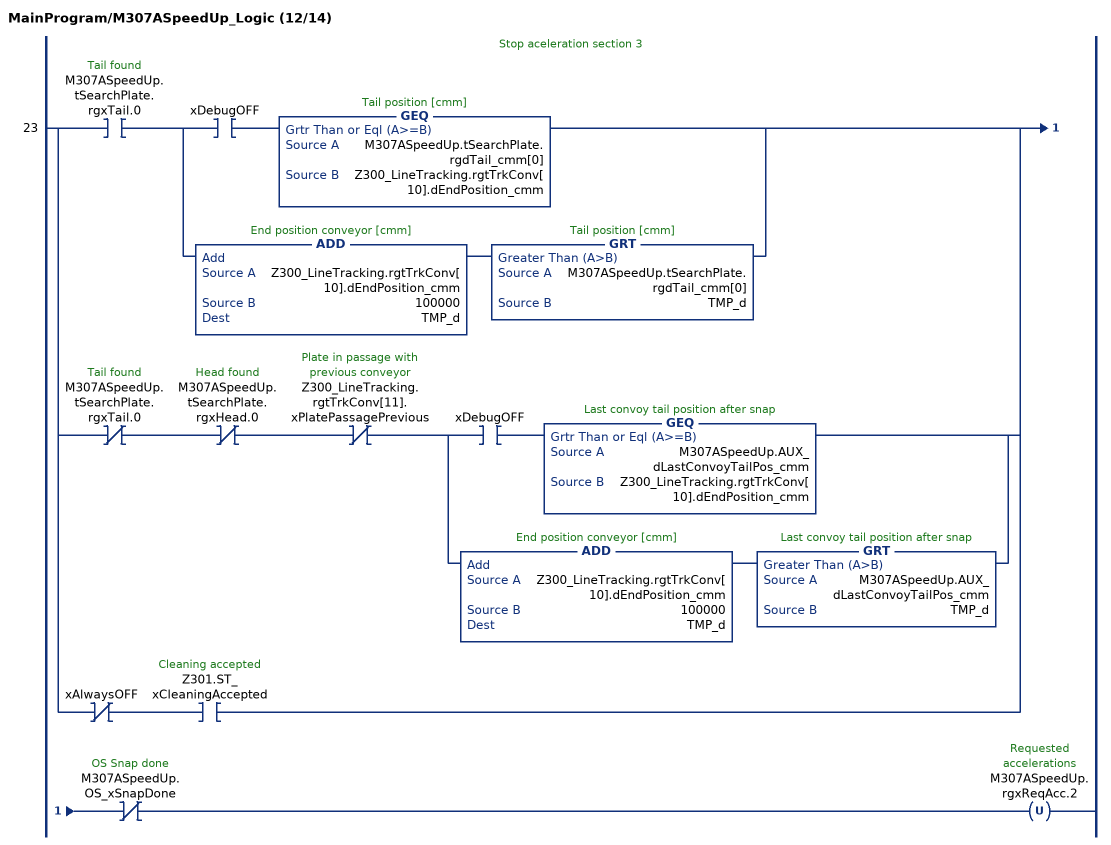
   // Stop aceleration section 3
   23: [XIC(M307ASpeedUp.tSearchPlate.rgxTail.0) [XIC(xDebugOFF) GEQ(M307ASpeedUp.tSearchPlate.rgdTail_cmm[0],Z300_LineTracking.rgtTrkConv[10].dEndPosition_cmm) ,ADD(Z300_LineTracking.rgtTrkConv[10].dEndPosition_cmm,100000,TMP_d) GRT(M307ASpeedUp.tSearchPlate.rgdTail_cmm[0],TMP_d) ] ,XIO(M307ASpeedUp.tSearchPlate.rgxTail.0) XIO(M307ASpeedUp.tSearchPlate.rgxHead.0) XIO(Z300_LineTracking.rgtTrkConv[11].xPlatePassagePrevious) [XIC(xDebugOFF) GEQ(M307ASpeedUp.AUX_dLastConvoyTailPos_cmm,Z300_LineTracking.rgtTrkConv[10].dEndPosition_cmm) ,ADD(Z300_LineTracking.rgtTrkConv[10].dEndPosition_cmm,100000,TMP_d) GRT(M307ASpeedUp.AUX_dLastConvoyTailPos_cmm,TMP_d) ] ,XIO(xAlwaysOFF) XIC(Z301.ST_xCleaningAccepted) ]XIO(M307ASpeedUp.OS_xSnapDone)OTU(M307ASpeedUp.rgxReqAcc.2);
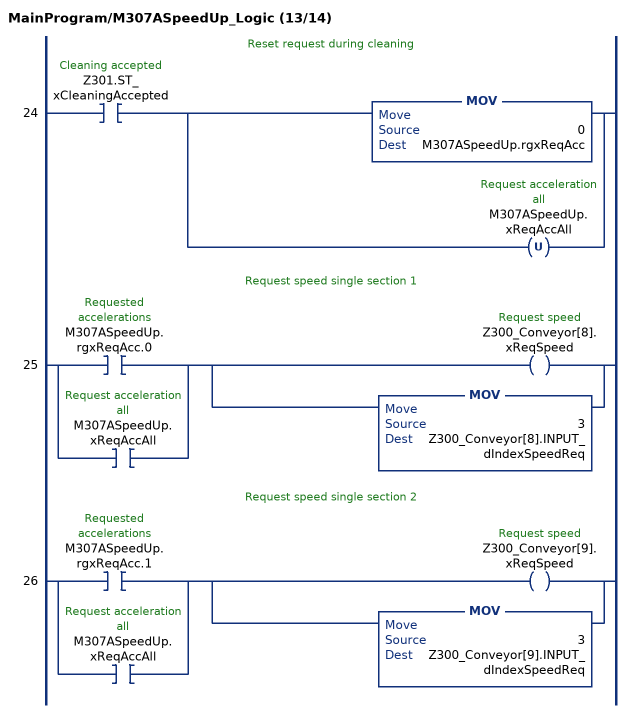
   // Reset request during cleaning
   24: XIC(Z301.ST_xCleaningAccepted)[MOV(0,M307ASpeedUp.rgxReqAcc) ,OTU(M307ASpeedUp.xReqAccAll) ];
   // Request speed single section 1
   25: [XIC(M307ASpeedUp.rgxReqAcc.0) ,XIC(M307ASpeedUp.xReqAccAll) ][OTE(Z300_Conveyor[8].xReqSpeed) ,MOV(3,Z300_Conveyor[8].INPUT_dIndexSpeedReq) ];
   // Request speed single section 2
   26: [XIC(M307ASpeedUp.rgxReqAcc.1) ,XIC(M307ASpeedUp.xReqAccAll) ][OTE(Z300_Conveyor[9].xReqSpeed) ,MOV(3,Z300_Conveyor[9].INPUT_dIndexSpeedReq) ];
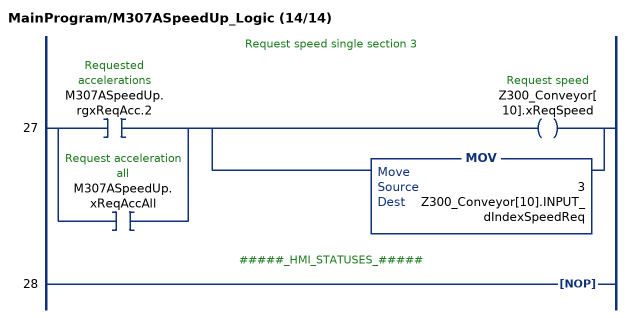
   // Request speed single section 3
   27: [XIC(M307ASpeedUp.rgxReqAcc.2) ,XIC(M307ASpeedUp.xReqAccAll) ][OTE(Z300_Conveyor[10].xReqSpeed) ,MOV(3,Z300_Conveyor[10].INPUT_dIndexSpeedReq) ];
   // #####_HMI_STATUSES_#####
   28: NOP();
END_ROUTINE

ROUTINE M30xTrimDeck_Faults   (* ladder *)
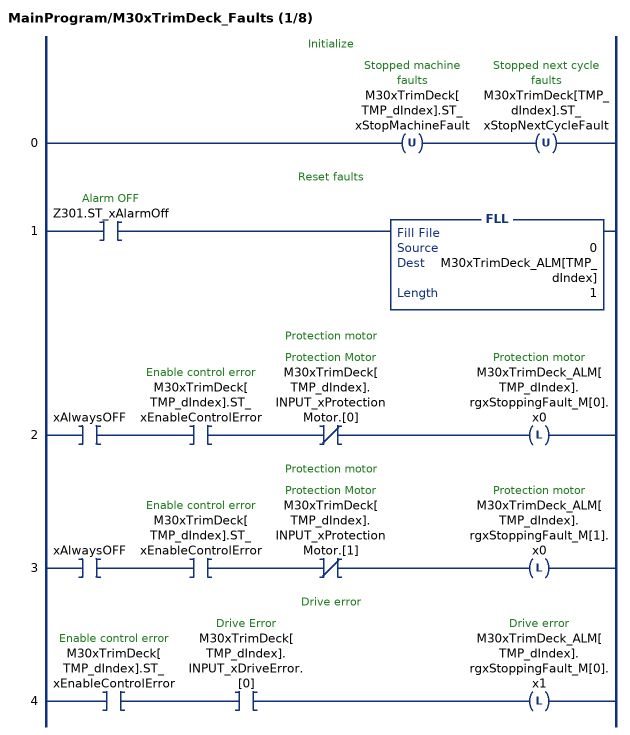
   // Initialize
   0: OTU(M30xTrimDeck[TMP_dIndex].ST_xStopMachineFault)OTU(M30xTrimDeck[TMP_dIndex].ST_xStopNextCycleFault);
   // Reset faults
   1: XIC(Z301.ST_xAlarmOff)FLL(0,M30xTrimDeck_ALM[TMP_dIndex],1);
   // Protection motor
   2: XIC(xAlwaysOFF)XIC(M30xTrimDeck[TMP_dIndex].ST_xEnableControlError)XIO(M30xTrimDeck[TMP_dIndex].INPUT_xProtectionMotor.[0])OTL(M30xTrimDeck_ALM[TMP_dIndex].rgxStoppingFault_M[0].x0);
   // Protection motor
   3: XIC(xAlwaysOFF)XIC(M30xTrimDeck[TMP_dIndex].ST_xEnableControlError)XIO(M30xTrimDeck[TMP_dIndex].INPUT_xProtectionMotor.[1])OTL(M30xTrimDeck_ALM[TMP_dIndex].rgxStoppingFault_M[1].x0);
   // Drive error
   4: XIC(M30xTrimDeck[TMP_dIndex].ST_xEnableControlError)XIC(M30xTrimDeck[TMP_dIndex].INPUT_xDriveError.[0])OTL(M30xTrimDeck_ALM[TMP_dIndex].rgxStoppingFault_M[0].x1);
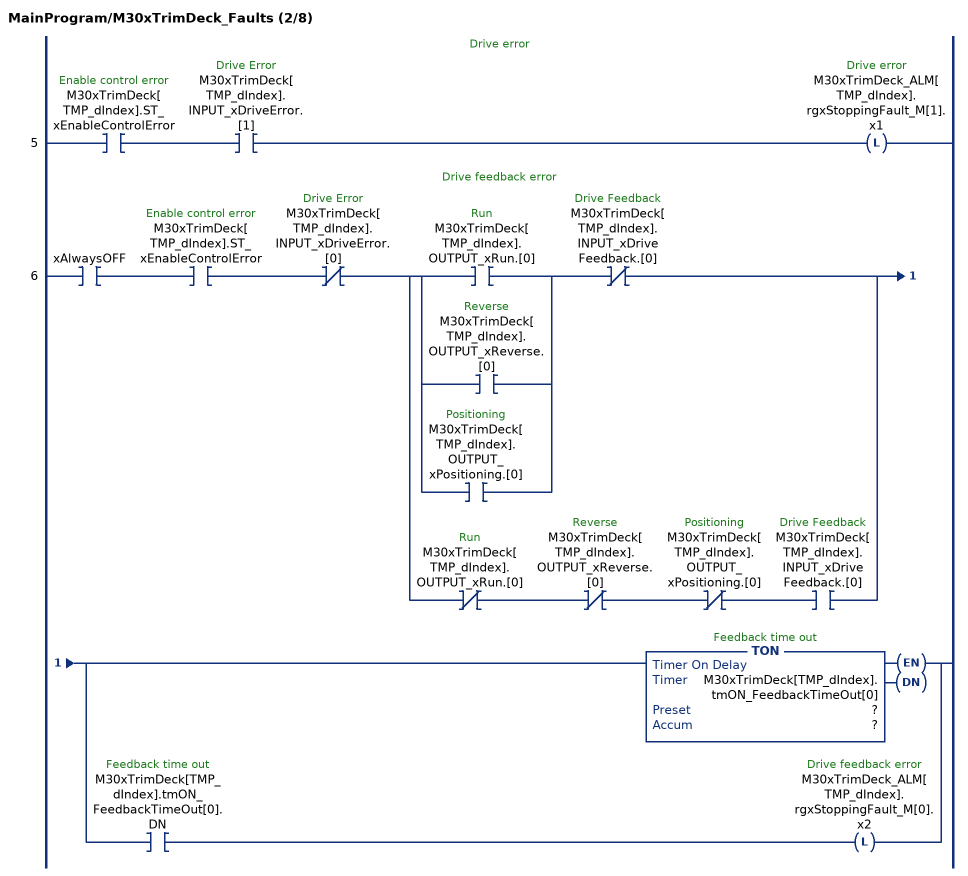
   // Drive error
   5: XIC(M30xTrimDeck[TMP_dIndex].ST_xEnableControlError)XIC(M30xTrimDeck[TMP_dIndex].INPUT_xDriveError.[1])OTL(M30xTrimDeck_ALM[TMP_dIndex].rgxStoppingFault_M[1].x1);
   // Drive feedback error
   6: XIC(xAlwaysOFF)XIC(M30xTrimDeck[TMP_dIndex].ST_xEnableControlError)XIO(M30xTrimDeck[TMP_dIndex].INPUT_xDriveError.[0])[[XIC(M30xTrimDeck[TMP_dIndex].OUTPUT_xRun.[0]) ,XIC(M30xTrimDeck[TMP_dIndex].OUTPUT_xReverse.[0]) ,XIC(M30xTrimDeck[TMP_dIndex].OUTPUT_xPositioning.[0]) ] XIO(M30xTrimDeck[TMP_dIndex].INPUT_xDriveFeedback.[0]) ,XIO(M30xTrimDeck[TMP_dIndex].OUTPUT_xRun.[0]) XIO(M30xTrimDeck[TMP_dIndex].OUTPUT_xReverse.[0]) XIO(M30xTrimDeck[TMP_dIndex].OUTPUT_xPositioning.[0]) XIC(M30xTrimDeck[TMP_dIndex].INPUT_xDriveFeedback.[0]) ][TON(M30xTrimDeck[TMP_dIndex].tmON_FeedbackTimeOut[0],?,?) ,XIC(M30xTrimDeck[TMP_dIndex].tmON_FeedbackTimeOut[0].DN) OTL(M30xTrimDeck_ALM[TMP_dIndex].rgxStoppingFault_M[0].x2) ];
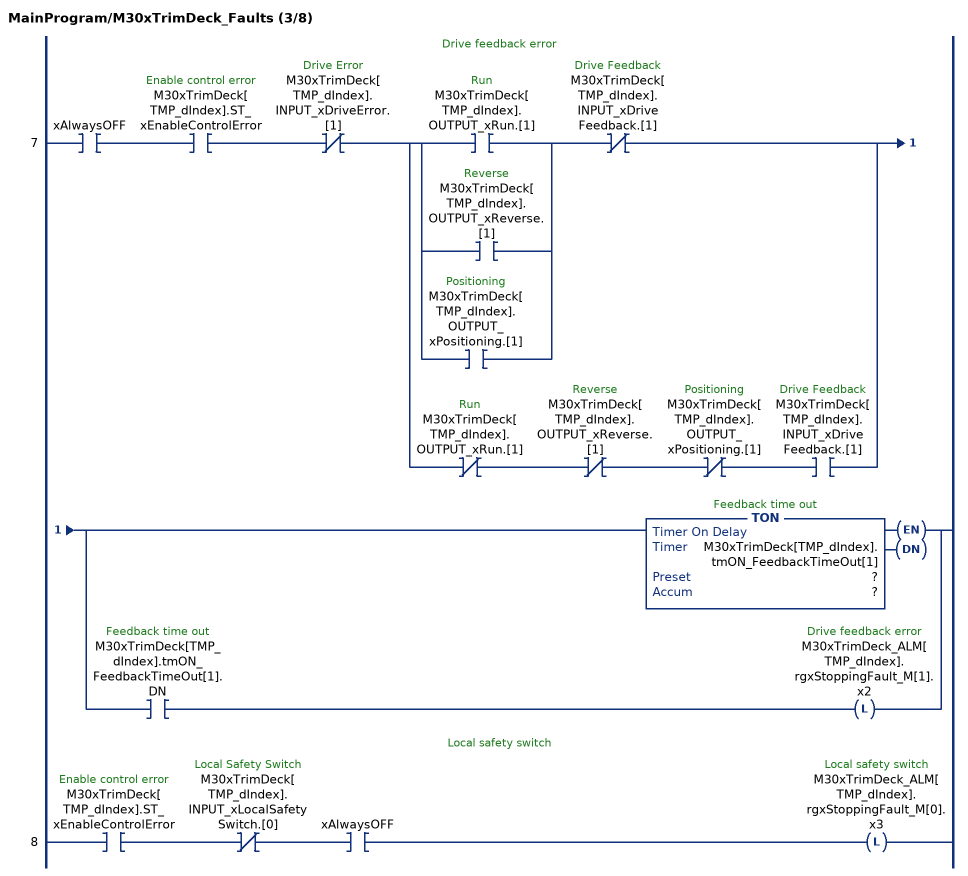
   // Drive feedback error
   7: XIC(xAlwaysOFF)XIC(M30xTrimDeck[TMP_dIndex].ST_xEnableControlError)XIO(M30xTrimDeck[TMP_dIndex].INPUT_xDriveError.[1])[[XIC(M30xTrimDeck[TMP_dIndex].OUTPUT_xRun.[1]) ,XIC(M30xTrimDeck[TMP_dIndex].OUTPUT_xReverse.[1]) ,XIC(M30xTrimDeck[TMP_dIndex].OUTPUT_xPositioning.[1]) ] XIO(M30xTrimDeck[TMP_dIndex].INPUT_xDriveFeedback.[1]) ,XIO(M30xTrimDeck[TMP_dIndex].OUTPUT_xRun.[1]) XIO(M30xTrimDeck[TMP_dIndex].OUTPUT_xReverse.[1]) XIO(M30xTrimDeck[TMP_dIndex].OUTPUT_xPositioning.[1]) XIC(M30xTrimDeck[TMP_dIndex].INPUT_xDriveFeedback.[1]) ][TON(M30xTrimDeck[TMP_dIndex].tmON_FeedbackTimeOut[1],?,?) ,XIC(M30xTrimDeck[TMP_dIndex].tmON_FeedbackTimeOut[1].DN) OTL(M30xTrimDeck_ALM[TMP_dIndex].rgxStoppingFault_M[1].x2) ];
   // Local safety switch
   8: XIC(M30xTrimDeck[TMP_dIndex].ST_xEnableControlError)XIO(M30xTrimDeck[TMP_dIndex].INPUT_xLocalSafetySwitch.[0])XIC(xAlwaysOFF)OTL(M30xTrimDeck_ALM[TMP_dIndex].rgxStoppingFault_M[0].x3);
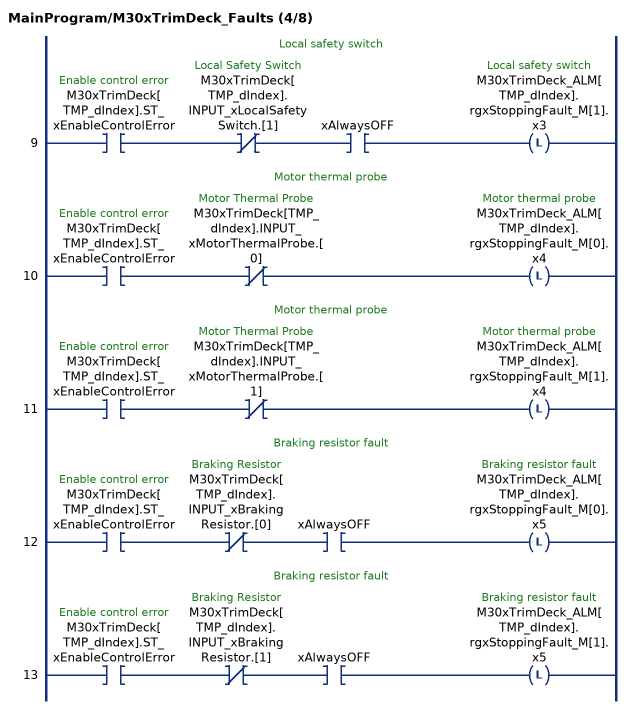
   // Local safety switch
   9: XIC(M30xTrimDeck[TMP_dIndex].ST_xEnableControlError)XIO(M30xTrimDeck[TMP_dIndex].INPUT_xLocalSafetySwitch.[1])XIC(xAlwaysOFF)OTL(M30xTrimDeck_ALM[TMP_dIndex].rgxStoppingFault_M[1].x3);
   // Motor thermal probe
   10: XIC(M30xTrimDeck[TMP_dIndex].ST_xEnableControlError)XIO(M30xTrimDeck[TMP_dIndex].INPUT_xMotorThermalProbe.[0])OTL(M30xTrimDeck_ALM[TMP_dIndex].rgxStoppingFault_M[0].x4);
   // Motor thermal probe
   11: XIC(M30xTrimDeck[TMP_dIndex].ST_xEnableControlError)XIO(M30xTrimDeck[TMP_dIndex].INPUT_xMotorThermalProbe.[1])OTL(M30xTrimDeck_ALM[TMP_dIndex].rgxStoppingFault_M[1].x4);
   // Braking resistor fault
   12: XIC(M30xTrimDeck[TMP_dIndex].ST_xEnableControlError)XIO(M30xTrimDeck[TMP_dIndex].INPUT_xBrakingResistor.[0])XIC(xAlwaysOFF)OTL(M30xTrimDeck_ALM[TMP_dIndex].rgxStoppingFault_M[0].x5);
   // Braking resistor fault
   13: XIC(M30xTrimDeck[TMP_dIndex].ST_xEnableControlError)XIO(M30xTrimDeck[TMP_dIndex].INPUT_xBrakingResistor.[1])XIC(xAlwaysOFF)OTL(M30xTrimDeck_ALM[TMP_dIndex].rgxStoppingFault_M[1].x5);
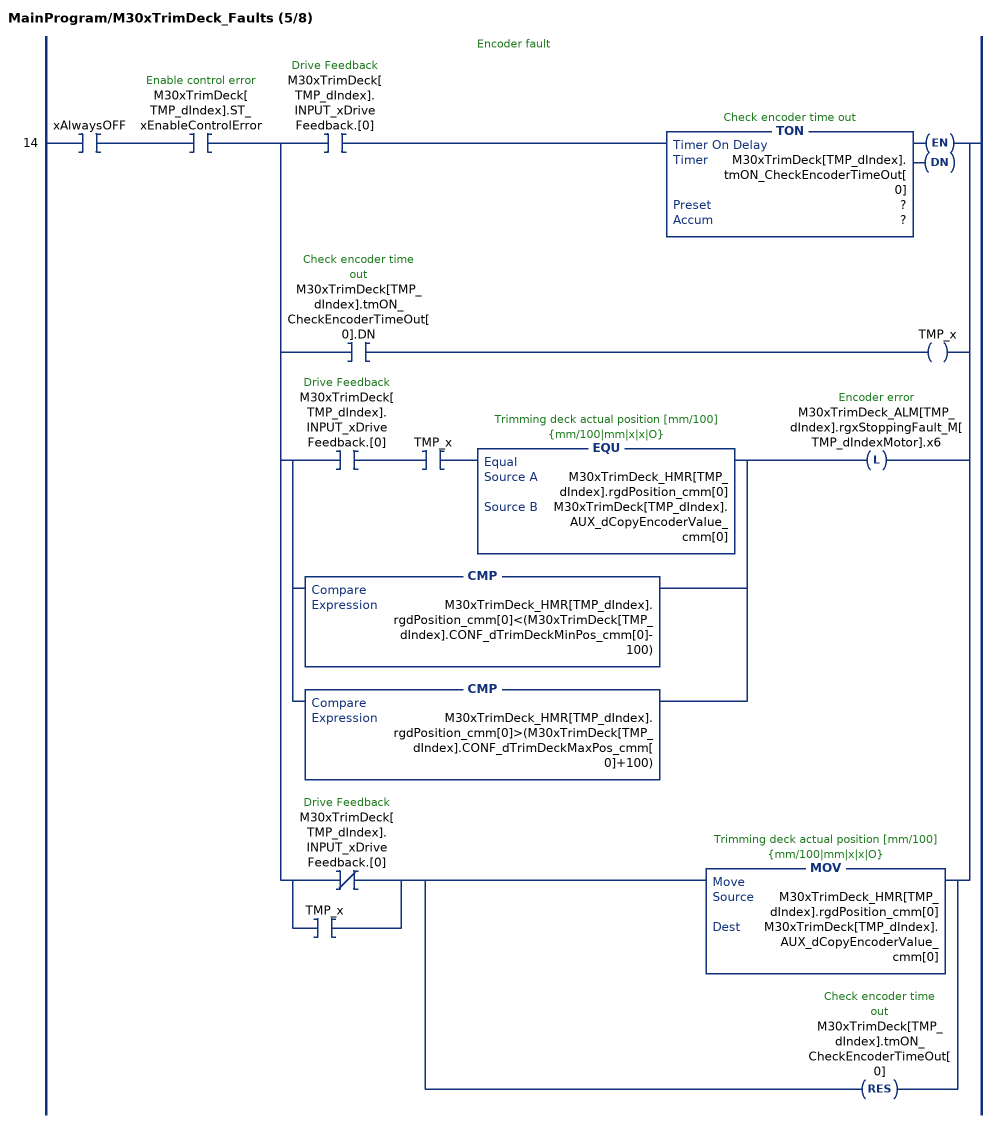
   // Encoder fault
   14: XIC(xAlwaysOFF)XIC(M30xTrimDeck[TMP_dIndex].ST_xEnableControlError)[XIC(M30xTrimDeck[TMP_dIndex].INPUT_xDriveFeedback.[0]) TON(M30xTrimDeck[TMP_dIndex].tmON_CheckEncoderTimeOut[0],?,?) ,XIC(M30xTrimDeck[TMP_dIndex].tmON_CheckEncoderTimeOut[0].DN) OTE(TMP_x) ,[XIC(M30xTrimDeck[TMP_dIndex].INPUT_xDriveFeedback.[0]) XIC(TMP_x) EQU(M30xTrimDeck_HMR[TMP_dIndex].rgdPosition_cmm[0],M30xTrimDeck[TMP_dIndex].AUX_dCopyEncoderValue_cmm[0]) ,CMP(M30xTrimDeck_HMR[TMP_dIndex].rgdPosition_cmm[0]<(M30xTrimDeck[TMP_dIndex].CONF_dTrimDeckMinPos_cmm[0]-100)) ,CMP(M30xTrimDeck_HMR[TMP_dIndex].rgdPosition_cmm[0]>(M30xTrimDeck[TMP_dIndex].CONF_dTrimDeckMaxPos_cmm[0]+100)) ] OTL(M30xTrimDeck_ALM[TMP_dIndex].rgxStoppingFault_M[TMP_dIndexMotor].x6) ,[XIO(M30xTrimDeck[TMP_dIndex].INPUT_xDriveFeedback.[0]) ,XIC(TMP_x) ] [MOV(M30xTrimDeck_HMR[TMP_dIndex].rgdPosition_cmm[0],M30xTrimDeck[TMP_dIndex].AUX_dCopyEncoderValue_cmm[0]) ,RES(M30xTrimDeck[TMP_dIndex].tmON_CheckEncoderTimeOut[0]) ] ];
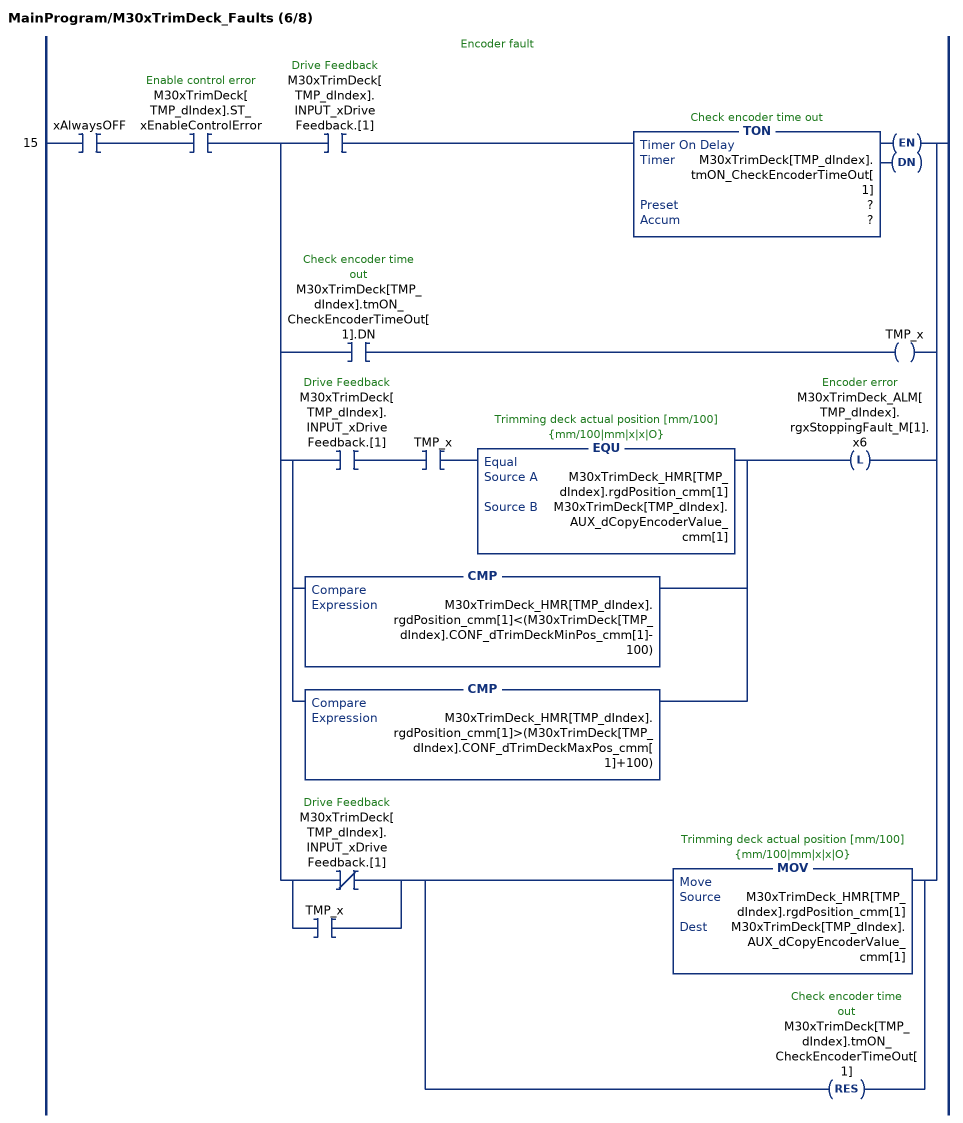
   // Encoder fault
   15: XIC(xAlwaysOFF)XIC(M30xTrimDeck[TMP_dIndex].ST_xEnableControlError)[XIC(M30xTrimDeck[TMP_dIndex].INPUT_xDriveFeedback.[1]) TON(M30xTrimDeck[TMP_dIndex].tmON_CheckEncoderTimeOut[1],?,?) ,XIC(M30xTrimDeck[TMP_dIndex].tmON_CheckEncoderTimeOut[1].DN) OTE(TMP_x) ,[XIC(M30xTrimDeck[TMP_dIndex].INPUT_xDriveFeedback.[1]) XIC(TMP_x) EQU(M30xTrimDeck_HMR[TMP_dIndex].rgdPosition_cmm[1],M30xTrimDeck[TMP_dIndex].AUX_dCopyEncoderValue_cmm[1]) ,CMP(M30xTrimDeck_HMR[TMP_dIndex].rgdPosition_cmm[1]<(M30xTrimDeck[TMP_dIndex].CONF_dTrimDeckMinPos_cmm[1]-100)) ,CMP(M30xTrimDeck_HMR[TMP_dIndex].rgdPosition_cmm[1]>(M30xTrimDeck[TMP_dIndex].CONF_dTrimDeckMaxPos_cmm[1]+100)) ] OTL(M30xTrimDeck_ALM[TMP_dIndex].rgxStoppingFault_M[1].x6) ,[XIO(M30xTrimDeck[TMP_dIndex].INPUT_xDriveFeedback.[1]) ,XIC(TMP_x) ] [MOV(M30xTrimDeck_HMR[TMP_dIndex].rgdPosition_cmm[1],M30xTrimDeck[TMP_dIndex].AUX_dCopyEncoderValue_cmm[1]) ,RES(M30xTrimDeck[TMP_dIndex].tmON_CheckEncoderTimeOut[1]) ] ];
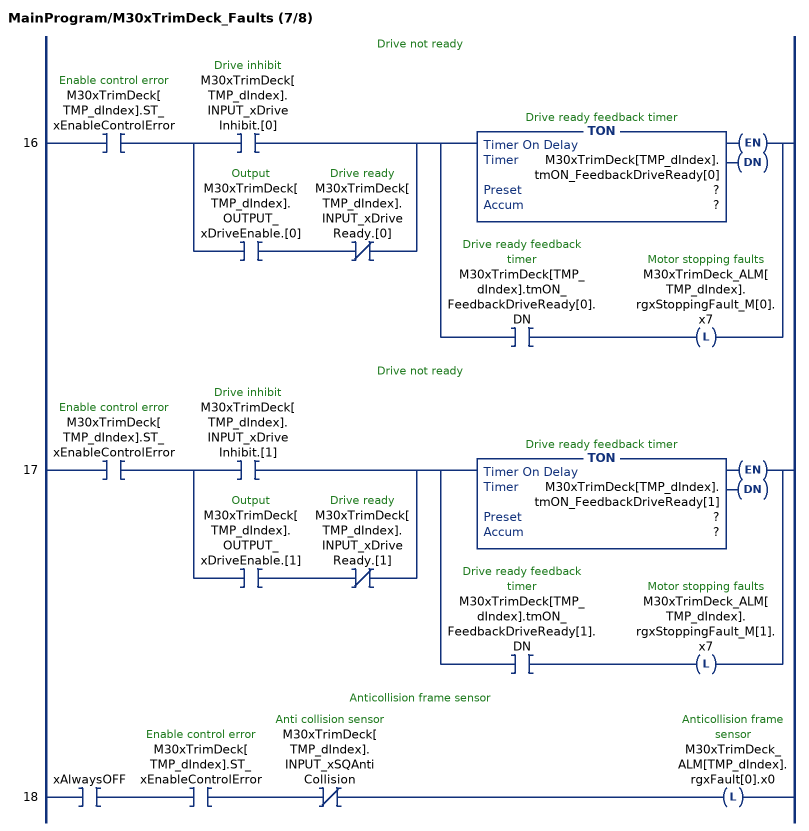
   // Drive not ready
   16: XIC(M30xTrimDeck[TMP_dIndex].ST_xEnableControlError)[XIC(M30xTrimDeck[TMP_dIndex].INPUT_xDriveInhibit.[0]) ,XIC(M30xTrimDeck[TMP_dIndex].OUTPUT_xDriveEnable.[0]) XIO(M30xTrimDeck[TMP_dIndex].INPUT_xDriveReady.[0]) ][TON(M30xTrimDeck[TMP_dIndex].tmON_FeedbackDriveReady[0],?,?) ,XIC(M30xTrimDeck[TMP_dIndex].tmON_FeedbackDriveReady[0].DN) OTL(M30xTrimDeck_ALM[TMP_dIndex].rgxStoppingFault_M[0].x7) ];
   // Drive not ready
   17: XIC(M30xTrimDeck[TMP_dIndex].ST_xEnableControlError)[XIC(M30xTrimDeck[TMP_dIndex].INPUT_xDriveInhibit.[1]) ,XIC(M30xTrimDeck[TMP_dIndex].OUTPUT_xDriveEnable.[1]) XIO(M30xTrimDeck[TMP_dIndex].INPUT_xDriveReady.[1]) ][TON(M30xTrimDeck[TMP_dIndex].tmON_FeedbackDriveReady[1],?,?) ,XIC(M30xTrimDeck[TMP_dIndex].tmON_FeedbackDriveReady[1].DN) OTL(M30xTrimDeck_ALM[TMP_dIndex].rgxStoppingFault_M[1].x7) ];
   // Anticollision frame sensor
   18: XIC(xAlwaysOFF)XIC(M30xTrimDeck[TMP_dIndex].ST_xEnableControlError)XIO(M30xTrimDeck[TMP_dIndex].INPUT_xSQAntiCollision)OTL(M30xTrimDeck_ALM[TMP_dIndex].rgxFault[0].x0);
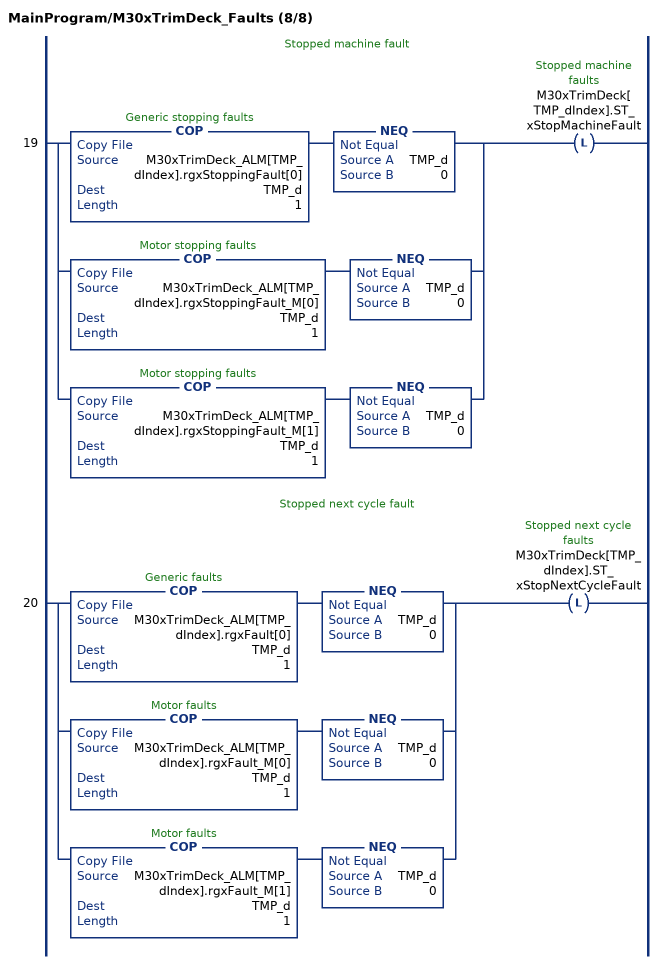
   // Stopped machine fault
   19: [COP(M30xTrimDeck_ALM[TMP_dIndex].rgxStoppingFault[0],TMP_d,1) NEQ(TMP_d,0) ,COP(M30xTrimDeck_ALM[TMP_dIndex].rgxStoppingFault_M[0],TMP_d,1) NEQ(TMP_d,0) ,COP(M30xTrimDeck_ALM[TMP_dIndex].rgxStoppingFault_M[1],TMP_d,1) NEQ(TMP_d,0) ]OTL(M30xTrimDeck[TMP_dIndex].ST_xStopMachineFault);
   // Stopped next cycle fault
   20: [COP(M30xTrimDeck_ALM[TMP_dIndex].rgxFault[0],TMP_d,1) NEQ(TMP_d,0) ,COP(M30xTrimDeck_ALM[TMP_dIndex].rgxFault_M[0],TMP_d,1) NEQ(TMP_d,0) ,COP(M30xTrimDeck_ALM[TMP_dIndex].rgxFault_M[1],TMP_d,1) NEQ(TMP_d,0) ]OTL(M30xTrimDeck[TMP_dIndex].ST_xStopNextCycleFault);
END_ROUTINE
